VERSION : 0.1
   VAR_IN_OUT
      commands : "Linked List: Method Interface: Search";
      list : "Linked List: List";
   END_VAR
   VAR_TEMP
      clear_commands : "Linked List: Method Interface: Search";
      found : Bool;
      pointer_list : DInt;
   END_VAR
   VAR CONSTANT
      no_error : String := 'no error';
      searched_empty_list : String := 'searched empty list';
   END_VAR
BEGIN
   REGION "EXIT CONDITION: SEARCHED EMPTY LIST"
       IF "Linked List: Private: Is Empty"(#list) THEN
           #commands := #clear_commands;
           #commands.out.not_found := TRUE;
           #commands.out.error := TRUE;
           #commands.out.error_message := #searched_empty_list;
           RETURN;
       END_IF;
   END_REGION

   REGION "SEARCH"
       FOR #pointer_list := 0 TO "LINKED_LIST_LENGTH" DO
           IF #list.me[#pointer_list].data = #commands.in.data THEN
               #found := TRUE;
               EXIT;
           END_IF;
       END_FOR;
   END_REGION

   REGION "FOUND"
       IF #found THEN
           #commands := #clear_commands;
           #commands.out.done := TRUE;
           #commands.out.found := TRUE;
           #commands.out.returned_node := #list.me[#pointer_list];
           #commands.out.error_message := #no_error;
           RETURN;
       END_IF;
   END_REGION

   REGION "NOT FOUND"
       IF NOT #found THEN
           #commands := #clear_commands;
           #commands.out.done := TRUE;
           #commands.out.not_found := TRUE;
           RETURN;
       END_IF;
   END_REGION
END_FUNCTION

FUNCTION "Linked List: Display" : Void   // FC172, SCL
{ S7_Optimized_Access := 'TRUE' }
VERSION : 0.1
   VAR_IN_OUT
      commands : "Linked List: Method Interface: Display";
      list : "Linked List: List";
   END_VAR
   VAR_TEMP
      clear_commands : "Linked List: Method Interface: Display";
   END_VAR
BEGIN
   #commands := #clear_commands;
   #commands.out.list := #list;
   #commands.out.done := TRUE;
END_FUNCTION

FUNCTION "Linked List: Insert" : Void   // FC173, SCL
{ S7_Optimized_Access := 'TRUE' }
VERSION : 0.1
   VAR_INPUT
      terminal_behavior : String;
   END_VAR
   VAR_IN_OUT
      commands : "Linked List: Method Interface: Insert";
      list : "Linked List: List";
   END_VAR
   VAR_TEMP
      clear_commands : "Linked List: Method Interface: Insert";
      current : "Linked List: Node";
      next_empty_node_index : DInt;
      previous : "Linked List: Node";
      next : "Linked List: Node";
   END_VAR
   VAR CONSTANT
      no_error : String := 'no error';
      inserted_into_full : String := 'attempted to insert into full list. delete a node and try again.';
      appended_as_head : String := 'appended as head of list';
   END_VAR
BEGIN
   REGION "EXIT CONDITION: INSERTED INTO FULL LIST"
       IF "Linked List: Private: Is Full"(#list) THEN
           #commands := #clear_commands;
           #commands.out.error := TRUE;
           #commands.out.error_message := #inserted_into_full;
           RETURN;
       END_IF;
   END_REGION

   REGION "EXIT CONDITION: INSERTED INTO EMPTY LIST"
       IF "Linked List: Private: Is Empty"(#list) THEN
           "Linked List: Private: Head an Empty List"(data := #commands.in.data,
                                                      terminal_behavior := #terminal_behavior,
                                                      list := #list);
           #commands := #clear_commands;
           #commands.out.error := TRUE;
           #commands.out.error_message := #appended_as_head;
           RETURN;
       END_IF;
   END_REGION

   REGION "GET INDEX OF NEXT EMPTY NODE"
       #next_empty_node_index := "Linked List: Private: Next Empty Node"(#list);
   END_REGION

   REGION "PREVIOUS, CURRENT, AND NEXT NODES"
       #current := #commands.in.target_node;
       #previous := "Linked List: Private: Get Previous"(current := #current,
                                                         list := #list);
       #next := #current;
   END_REGION

   REGION "INSERT BEFORE TARGET NODE"
       // new node's data becomes command data
       #list.me[#next_empty_node_index].data := #commands.in.data;
       // new node's key becomes array index
       #list.me[#next_empty_node_index].meta.key := #next_empty_node_index;
       // shorten name for indexing
       #current := #list.me[#next_empty_node_index];
       // insert
       IF NOT #next.meta.is_head THEN
           "Linked List: Private: After"(node := #list.me[#current.meta.key],
                                         previous_node := #list.me[#previous.meta.key]);
       END_IF;
       "Linked List: Private: Before"(next_node := #list.me[#next.meta.key],
                                      node := #list.me[#current.meta.key]);
   END_REGION

   REGION "COMMANDS OUT"
       #commands := #clear_commands;
       #commands.out.done := TRUE;
       #commands.out.error_message := #no_error;
   END_REGION
END_FUNCTION

FUNCTION "Linked List: Reverse" : Void   // FC174, SCL
{ S7_Optimized_Access := 'TRUE' }
VERSION : 0.1
   VAR_IN_OUT
      commands : "Linked List: Method Interface: Reverse";
      list : "Linked List: List";
   END_VAR
   VAR_TEMP
      clear_commands : "Linked List: Method Interface: Reverse";
      current : "Linked List: Node";
      next : "Linked List: Node";
      previous : "Linked List: Node";
      null_node : "Linked List: Node";
   END_VAR
   VAR CONSTANT
      no_error : String := 'no error';
      reversed_empty_list : String := 'reversed empty list';
   END_VAR
BEGIN
   IF "Linked List: Private: Is Empty"(#list) THEN
       #commands := #clear_commands;
       #commands.out.error := TRUE;
       #commands.out.error_message := #reversed_empty_list;
       RETURN;
   END_IF;

   "Linked List: Private: Clear Node"(#null_node);
   #previous := #null_node;
   #current := "Linked List: Private: Get Head"(#list);
   #list.me[#current.meta.key].meta.is_head := FALSE;
   #list.me[#current.meta.key].meta.is_tail := TRUE;
   WHILE #current.meta.next <> "NULL_TOKEN" DO
       #next := #list.me[#current.meta.next];
       #list.me[#current.meta.key].meta.next := #previous.meta.key;
       #previous := #current;
       #current := #next;
       #list.me[#current.meta.key].meta.is_head := FALSE;
       #list.me[#current.meta.key].meta.is_tail := FALSE;
   END_WHILE;
   #list.me[#current.meta.key].meta.next := #previous.meta.key;
   #list.me[#current.meta.key].meta.is_head := TRUE;
   #list.me[#current.meta.key].meta.is_tail := FALSE;

   #commands := #clear_commands;
   #commands.out.done := TRUE;
   #commands.out.error_message := #no_error;
END_FUNCTION

FUNCTION "Linked List: Reset" : Void   // FC175, SCL
{ S7_Optimized_Access := 'TRUE' }
VERSION : 0.1
   VAR_IN_OUT
      commands : "Linked List: Method Interface: Reset";
      list : "Linked List: List";
   END_VAR
   VAR_TEMP
      blank_node : "Linked List: Node";
      list_pointer : DInt;
      clear_commands : "Linked List: Method Interface: Reset";
   END_VAR
BEGIN
   FOR #list_pointer := 0 TO "LINKED_LIST_LENGTH" DO
       "Linked List: Private: Clear Node"(#list.me[#list_pointer]);
   END_FOR;
   #commands := #clear_commands;
   #commands.out.done := TRUE;
END_FUNCTION

// folder: OBs

ORGANIZATION_BLOCK "Rack or station failure"   // OB86, LAD, RackStationFailure
{ S7_Optimized_Access := 'TRUE' }
VERSION : 0.1
   VAR_INPUT
      LADDR : Hw_Device;   // Hardware identifier
      Event_Class : Byte;   // Event class
      Fault_ID : Byte;   // Fault identifier
   END_VAR
BEGIN
END_ORGANIZATION_BLOCK

ORGANIZATION_BLOCK "Startup"   // OB100, LAD, Startup
TITLE = "Complete Restart"
{ S7_Optimized_Access := 'TRUE' }
VERSION : 0.1
   VAR_INPUT
      LostRetentive : Bool;   // True if retentive data are lost
      LostRTC : Bool;   // True if date and time are lost
   END_VAR
   VAR CONSTANT
      ALLOTTED : Real := 1800.0;
      CRITICAL : Real := 300.0;
   END_VAR
BEGIN

REGION Network 1
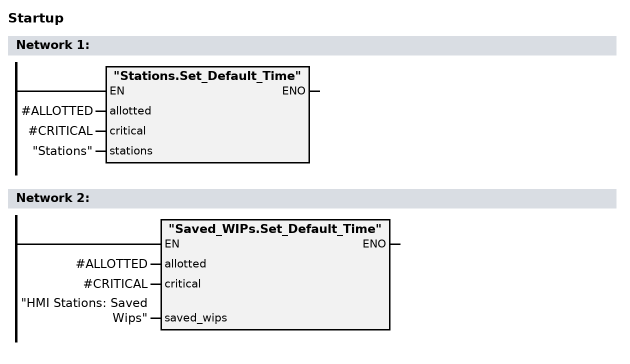
   RUNG wire#powerrail
      "Stations.Set_Default_Time"(allotted := #ALLOTTED, critical := #CRITICAL, stations := "Stations")
   END_RUNG
   // the same network as SCL:
   "Stations.Set_Default_Time"(allotted := #ALLOTTED, critical := #CRITICAL, stations := "Stations");
END_REGION

REGION Network 2
   RUNG wire#powerrail
      "Saved_WIPs.Set_Default_Time"(allotted := #ALLOTTED, critical := #CRITICAL, saved_wips := "HMI Stations: Saved Wips")
   END_RUNG
   // the same network as SCL:
   "Saved_WIPs.Set_Default_Time"(allotted := #ALLOTTED,
                           critical := #CRITICAL,
                           saved_wips := "HMI Stations: Saved Wips");
END_REGION
END_ORGANIZATION_BLOCK

ORGANIZATION_BLOCK "Programming error"   // OB121, LAD, ProgrammingError
{ S7_Optimized_Access := 'TRUE' }
VERSION : 0.1
   VAR_INPUT
      BlockNr : UInt;   // Number of causing block
      Reaction : USInt;   // 0:ignore, 1:substitute, 2:skip
      Fault_ID : Byte;   // Fault identifier
      BlockType : USInt;   // 16#01:OB, 16#02:FC, 16#03:FB, 16#04:SFC, 16#05:SFB, 16#06:DB: Type of block causing the error
      Area : USInt;   // Area where the error occured
      DBNr : DB_ANY;   // DB number if Area = DB or DI
      Csg_OBNr : OB_Any;   // Number of OB causing the error
      Csg_Prio : USInt;   // Priority of OB causing the error
      Width : USInt;   // 0:bit, 1:byte, 2:word, 3:dword, 4:lword
   END_VAR
BEGIN
END_ORGANIZATION_BLOCK

ORGANIZATION_BLOCK "IO access error"   // OB122, LAD, IOAccessError
{ S7_Optimized_Access := 'TRUE' }
VERSION : 0.1
   VAR_INPUT
      BlockNr : UInt;   // Number of causing block
      Reaction : USInt;   // 0:ignore, 1:substitute, 2:skip
      Fault_ID : Byte;   // 16#42:reading, 16#43:writing
      BlockType : USInt;   // 16#01:OB, 16#02:FC, 16#03:FB, 16#04:SFC, 16#05:SFB, 16#06:DB: Type of block causing the error
      Area : USInt;   // 16#81:I, 16#82:Q: IO area where the IOaccess error occured
      DBNr : DB_ANY;   // Reserved for system
      Csg_OBNr : OB_Any;   // Number of OB causing the error
      Csg_Prio : USInt;   // Priority of OB causing the error
      Width : USInt;   // 0:bit, 1:byte, 2:word, 3:dword, 4:lword
   END_VAR
BEGIN
END_ORGANIZATION_BLOCK

// folder: Order/States

FUNCTION_BLOCK "Order_State"   // FB2, SCL
{ S7_Optimized_Access := 'TRUE' }
VERSION : 0.1
   VAR_INPUT
      part_number_library : "Recipe: PN Text Library";
   END_VAR
   VAR_IN_OUT
      stations : "Station: All Stations";
   END_VAR
   VAR_TEMP
      station_pointer : Int;
      button_pointer : Int;
      station : "Station: Single Station";
   END_VAR
BEGIN
   REGION "FOR EACH STATION"
       FOR #station_pointer := 0 TO "STATION_COUNT" DO

           REGION "POPULATE CURRENT STATION"
               #station := #stations.stn[#station_pointer];
           END_REGION

           REGION "SET TO IDLE ON WIP SWAP"
               IF #station.flags.wipSwapped THEN
                   CONTINUE;
               END_IF;
           END_REGION

           REGION "FOR EACH BUTTON"
               FOR #button_pointer := 0 TO "BUTTON_COUNT" DO

                   REGION "INITIALIZE STATE"
                       "Order_State.Initialize_State"(newParams := #station.wipCmpts.flags.new_part_number,
                                                      pnGood := #station.wipCmpts.flags.part_number_good[#button_pointer],
                                                      state := #station.wipCmpts.orderState[#button_pointer]);
                   END_REGION

                   REGION "ENTER IDLE"
                       "Order_State.Enter_Idle"(part_button_falling_edge := #station.wipCmpts.kp8Logical.falling.btn[#button_pointer],
                                                state := #station.wipCmpts.orderState[#button_pointer]);
                   END_REGION

                   REGION "ENTER REQUESTED"
                       "Order_State.Enter_Requested"(btnRising := #station.wipCmpts.kp8Logical.rising.btn[#button_pointer],
                                                     state := #station.wipCmpts.orderState[#button_pointer]);
                   END_REGION

                   REGION "ENTER REQUESTED CRITICAL"
                       "Order_State.Enter_Requested_Critical"(timerVal := #station.wipCmpts.timers.remaining[#button_pointer],
                                                              state := #station.wipCmpts.orderState[#button_pointer]);
                   END_REGION

                   REGION "ENTER REQUESTED EXPIRED"
                       "Order_State.Enter_Requested_Expired"(timerVal := #station.wipCmpts.timers.remaining[#button_pointer],
                                                             state := #station.wipCmpts.orderState[#button_pointer]);
                   END_REGION

                   REGION "SAVE CURRENT STATION"
                       #stations.stn[#station_pointer] := #station;
                   END_REGION

               END_FOR;
           END_REGION

       END_FOR;
   END_REGION
END_FUNCTION_BLOCK

FUNCTION "Order_State.Enter_Idle" : Void   // FC6, SCL
{ S7_Optimized_Access := 'TRUE' }
VERSION : 0.1
   VAR_INPUT
      part_button_falling_edge : Bool;
   END_VAR
   VAR_IN_OUT
      state : Int;
   END_VAR
BEGIN
   IF #part_button_falling_edge THEN
       #state := "IDLE";
       RETURN;
   END_IF;
END_FUNCTION

FUNCTION "Order_State.Enter_Requested" : Void   // FC7, SCL
{ S7_Optimized_Access := 'TRUE' }
VERSION : 0.1
   VAR_INPUT
      btnRising : Bool;
   END_VAR
   VAR_IN_OUT
      state : Int;
   END_VAR
BEGIN
   IF #state = "IDLE" THEN
       IF #btnRising THEN
           #state := "REQUESTED";
       END_IF;
   END_IF;
END_FUNCTION

FUNCTION "Order_State.Initialize_State" : Void   // FC10, SCL
{ S7_Optimized_Access := 'TRUE' }
VERSION : 0.1
   VAR_INPUT
      newParams : Bool;
      pnGood : Bool;
   END_VAR
   VAR_IN_OUT
      state : Int;
   END_VAR
BEGIN
   REGION "ON NEW PARAMETERS"
       IF #newParams THEN
           #state := BOOL_TO_INT(#pnGood);
       END_IF;
   END_REGION
END_FUNCTION

FUNCTION "Order_State.Enter_Requested_Critical" : Void   // FC16, SCL
{ S7_Optimized_Access := 'TRUE' }
VERSION : 0.1
   VAR_INPUT
      timerVal : Real;
   END_VAR
   VAR_IN_OUT
      state : Int;
   END_VAR
   VAR_TEMP
      temp : Real;
   END_VAR
BEGIN
   IF #state = "REQUESTED" THEN
       IF #timerVal > 0.0 AND #timerVal <= "DEFAULT_CRITICAL_TIME" THEN
           #state := "REQUESTED_CRITICAL";
       END_IF;
   END_IF;
END_FUNCTION

FUNCTION "Order_State.Enter_Requested_Expired" : Void   // FC17, SCL
{ S7_Optimized_Access := 'TRUE' }
VERSION : 0.1
   VAR_INPUT
      timerVal : Real;
   END_VAR
   VAR_IN_OUT
      state : Int;
   END_VAR
BEGIN
   IF #state = "REQUESTED_CRITICAL" THEN
       IF #timerVal <= -0.001 THEN
           #state := "REQUESTED_EXPIRED";
       END_IF;
   END_IF;
END_FUNCTION

FUNCTION "Order_State.Enter_Ordered" : Void   // FC297, SCL
{ S7_Optimized_Access := 'TRUE' }
VERSION : 0.1
   VAR_INPUT
      address : DInt;
   END_VAR
   VAR_IN_OUT
      stations : "Station: All Stations";
   END_VAR
BEGIN
   "Order_State.Set_State_by_Address"(address := #address,
                                      state := "ORDERED",
                                      stations := #stations);
END_FUNCTION

FUNCTION "Order_State.Enter_Acknowledged" : Void   // FC301, SCL
{ S7_Optimized_Access := 'TRUE' }
VERSION : 0.1
   VAR_INPUT
      address : DInt;
   END_VAR
   VAR_IN_OUT
      stations : "Station: All Stations";
   END_VAR
BEGIN
   "Order_State.Set_State_by_Address"(address := #address,
                                      state := "ACKNOWLEGED",
                                      stations := #stations);
END_FUNCTION

FUNCTION "Order_State.Set_State_by_Address" : Void   // FC302, SCL
{ S7_Optimized_Access := 'TRUE' }
VERSION : 0.1
   VAR_INPUT
      address : DInt;
      state : Int;
   END_VAR
   VAR_IN_OUT
      stations : "Station: All Stations";
   END_VAR
   VAR_TEMP
      _p_button : DInt;
      _p_station : DInt;
      _p_wip : DInt;
   END_VAR
BEGIN
   #_p_button := "Address.Get_Button"(#address);
   #_p_station := "Address.Get_Station"(#address);
   #_p_wip := "Address.Get_Wip"(#address);
   #stations.stn[#_p_station].wipCmpts.orderState[#_p_button] := #state;
END_FUNCTION

FUNCTION "Order_State.Swap_WIP_States" : Void   // FC317, SCL
{ S7_Optimized_Access := 'TRUE' }
VERSION : 0.1
   VAR_IN_OUT
      station : "Station: Single Station";
   END_VAR
   VAR_TEMP
      _length : Int;
      _button_pointer : Int;
   END_VAR
BEGIN
   #_length := UDINT_TO_INT("Array.Any.Length"(#station.wipCmpts.pnCode)) - 1;
   FOR #_button_pointer := 0 TO #_length DO
       IF #station.wipCmpts.pnCode[#_button_pointer] <= 0 THEN
           #station.wipCmpts.orderState[#_button_pointer] := 0;
           CONTINUE;
       END_IF;
       IF #station.wipCmpts.orderState[#_button_pointer] <> 0 THEN
           CONTINUE;
       END_IF;
       #station.wipCmpts.orderState[#_button_pointer] := "IDLE";
   END_FOR;
END_FUNCTION

// folder: Order/Timers

FUNCTION_BLOCK "Order Timer"   // FB6, SCL
{ S7_Optimized_Access := 'TRUE' }
VERSION : 0.1
   VAR_INPUT
      pnLib : "Recipe: PN Text Library";
   END_VAR
   VAR_IN_OUT
      stns : "Station: All Stations";
   END_VAR
   VAR
      rt : "Runtime Data";
   END_VAR
   VAR_TEMP
      pStn : Int;
      pBtn : Int;
   END_VAR
BEGIN
   REGION "RUNTIME CALL"
       #rt.elapsed := RUNTIME(#rt.mem);
       #rt.asReal := LREAL_TO_REAL(#rt.elapsed);
   END_REGION

   REGION "FOR EACH STATION"
       FOR #pStn := 0 TO "STATION_COUNT" DO

           REGION "FOR EACH BUTTON"
               FOR #pBtn := 0 TO "BUTTON_COUNT" DO

                   REGION "INITIALIZE TIMERS"
                       "Order Timer: Initialize"(pnLib := #pnLib,
                                                 pBtn := #pBtn,
                                                 stn := #stns.stn[#pStn]);
                   END_REGION

                   REGION "EXECUTE TIMERS"
                       "Order Timer: Timer Execution"(elapsedTime := #rt.asReal,
                                                      pBtn := #pBtn,
                                                      stn:=#stns.stn[#pStn],
                                                      timers := #stns.stn[#pStn].wipCmpts.timers);
                   END_REGION

               END_FOR;
           END_REGION

       END_FOR;
   END_REGION
END_FUNCTION_BLOCK

FUNCTION "Order Timer: Initialize" : Void   // FC8, SCL
{ S7_Optimized_Access := 'TRUE' }
VERSION : 0.1
   VAR_INPUT
      pnLib : "Recipe: PN Text Library";
      pBtn : Int;
   END_VAR
   VAR_IN_OUT
      stn : "Station: Single Station";
   END_VAR
   VAR_TEMP
      pnGood : Bool;
      default : Bool;
      clear : Bool;
   END_VAR
BEGIN
   REGION "ON PN CHANGE"
       IF #stn.wipCmpts.flags.new_part_number THEN

           REGION "INITIALIZE TO DEFAULT"

               REGION "EXECUTION VALIDATION"
                   #default := "Order Timer: Set to Default Check"(pnGood := #stn.wipCmpts.flags.part_number_good[#pBtn],
                                                                   inSettingsScreen := #stn.wipCmpts.flags.in_settings_screen,
                                                                   timerReset := #stn.wipCmpts.flags.reset_timer[#pBtn]);
               END_REGION

               REGION "ON VALIDATION"
                   IF #default THEN

                       REGION "SET DEFAULT TIME VALUE"
                           #stn.wipCmpts.timers.ptAllotted[#pBtn] := "DEFAULT_TOTAL_TIME";
                           #stn.wipCmpts.timers.ptCritical[#pBtn] := "DEFAULT_CRITICAL_TIME";
                       END_REGION

                   END_IF;
               END_REGION

           END_REGION

           REGION "INITIALIZE TO ZERO"

               REGION "EXECUTION VALIDATION"
                   #clear := "Order Timer: Set to Zero Check"(pnGood := #stn.wipCmpts.flags.part_number_good[#pBtn],
                                                              inSettingsScreen := #stn.wipCmpts.flags.in_settings_screen,
                                                              timerReset := #stn.wipCmpts.flags.reset_timer[#pBtn]);
               END_REGION

               REGION "ON VALIDATION"
                   IF #clear THEN

                       REGION "SET DEFAULT TIME VALUE"
                           #stn.wipCmpts.timers.ptAllotted[#pBtn] := 0.0;
                           #stn.wipCmpts.timers.ptCritical[#pBtn] := 0.0;
                       END_REGION

                   END_IF;
               END_REGION

           END_REGION

       END_IF;
   END_REGION
END_FUNCTION

FUNCTION "Order Timer: Timer Execution" : Void   // FC11, SCL
{ S7_Optimized_Access := 'TRUE' }
VERSION : 0.1
   VAR_INPUT
      elapsedTime : Real;
      pBtn : Int;
      stn : "Station: Single Station";
   END_VAR
   VAR_IN_OUT
      timers : "Request_Timers.UDT";
   END_VAR
BEGIN
   REGION "RUN CONDITIONS"
       CASE #stn.wipCmpts.orderState[#pBtn] OF

           "RESET", "IDLE":
               IF #stn.flags.stateTransition[#pBtn] THEN
                   #timers.elapsed[#pBtn] := 0.0;
                   #timers.remaining[#pBtn] := 0.0;
               END_IF;

           "REQUESTED".."ACKNOWLEDGED_EXPIRED":
               #timers.elapsed[#pBtn] += #elapsedTime;
               #timers.remaining[#pBtn] := #timers.ptAllotted[#pBtn] - #timers.elapsed[#pBtn];

           ELSE:
               ;

       END_CASE;
   END_REGION
END_FUNCTION

FUNCTION "Order Timer: Set to Default Check" : Bool   // FC12, SCL
{ S7_Optimized_Access := 'TRUE' }
VERSION : 0.1
   VAR_INPUT
      pnGood : Bool;
      inSettingsScreen : Bool;
      timerReset : Bool;
   END_VAR
   VAR_TEMP
      ret : Bool;
   END_VAR
BEGIN
   REGION "ON VALID PN"
       #ret := #pnGood;
   END_REGION

   REGION "NOT WHILE IN SETTINGS SCREEN"
       IF #inSettingsScreen THEN
           #ret := FALSE;
       END_IF;
   END_REGION

   REGION "ON RESET REQUEST"
       #ret := #timerReset OR #ret;
   END_REGION

   REGION "RETURN"
       #"Order Timer: Set to Default Check" := #ret;
   END_REGION
END_FUNCTION

FUNCTION "Order Timer: Set to Zero Check" : Bool   // FC15, SCL
{ S7_Optimized_Access := 'TRUE' }
VERSION : 0.1
   VAR_INPUT
      pnGood : Bool;
      inSettingsScreen : Bool;
      timerReset : Bool;
   END_VAR
   VAR_TEMP
      ret : Bool;
   END_VAR
BEGIN
   REGION "ON VALID PN"
       #ret := NOT #pnGood;
   END_REGION

   REGION "NOT WHILE IN SETTINGS SCREEN"
       IF #inSettingsScreen THEN
           #ret := FALSE;
       END_IF;
   END_REGION

   REGION "ON RESET REQUEST"
       #ret := #timerReset OR #ret;
   END_REGION

   REGION "RETURN"
       #"Order Timer: Set to Zero Check" := #ret;
   END_REGION
END_FUNCTION

// folder: Part Request

FUNCTION_BLOCK "Part Request"   // FB7, SCL
{ S7_Optimized_Access := 'TRUE' }
VERSION : 0.1
   VAR_INPUT
      stns : "Station: All Stations";
      savedWips : "Recipe: HMI Stations Saved Wips";
      pnLib : "Recipe: PN Text Library";
   END_VAR
   VAR_IN_OUT
      dataTable : "Part Request Data";
   END_VAR
   VAR RETAIN
      pDataRow : Int;
   END_VAR
   VAR_TEMP
      address : DInt;
      addRequest : Bool;
      inTable : DInt;
      pStn : Int;
      pBtn : Int;
      pWip : Int;
      pRqstsRow : Int;
      removeRequest : Bool;
   END_VAR
BEGIN
   REGION "FOR EACH STATION"
       FOR #pStn := 0 TO "STATION_COUNT" DO

           REGION "FOR EACH BUTTON"
               FOR #pBtn := 0 TO "BUTTON_COUNT" DO

                   REGION "NEXT BUTTON ON NO TRANSITION"
                       IF NOT #stns.stn[#pStn].flags.stateTransition[#pBtn] THEN
                           CONTINUE;
                       END_IF;
                   END_REGION

                   REGION "GET ADDRESS"
                       #pWip := DINT_TO_INT(#stns.stn[#pStn].wipData.index);
                       #address := "Address.Set_Address"(pStn := #pStn, pBtn := #pBtn, pWip := #pWip);
                   END_REGION

                   REGION "CHECK FOR ENTRY IN DATA TABLE"
                       #inTable := "Part Request: Address in Table"(address := #address,
                                                                    table := #dataTable);
                   END_REGION

                   REGION "ADD"

                       REGION "VALIDATE CONDITIONS"
                           #addRequest := "Part Request: Validate Add"(inTable := #inTable,
                                                                       orderState := #stns.stn[#pStn].wipCmpts.orderState[#pBtn]);
                       END_REGION

                       REGION "EXECUTE"
                           IF #addRequest THEN
                               #addRequest := FALSE;
                               #dataTable.row[#pDataRow] := #address;
                               "Row Pointer: Roll Over"(limit := "partReqDataRowCount",
                                                        "pointer" := #pDataRow);
                           END_IF;
                       END_REGION

                   END_REGION

                   REGION "REMOVE SINGLE STATION"

                       REGION "VALIDATE CONDITIONS: SINGLE"
                           #removeRequest := "Part Request: Validate Remove: Single"(inTable := #inTable,
                                                                                     orderState := #stns.stn[#pStn].wipCmpts.orderState[#pBtn]);
                       END_REGION

                       REGION "EXECUTE"
                           IF #removeRequest THEN
                               #removeRequest := FALSE;
                               #dataTable.row[#inTable] := -1;
                               "Part Request: Collapse Table"(#dataTable);
                               "Row Pointer: Post Collapse"(dataTable := #dataTable,
                                                            pDataRow := #pDataRow);
                           END_IF;
                       END_REGION

                   END_REGION

               END_FOR;
           END_REGION

       END_FOR;
   END_REGION
END_FUNCTION_BLOCK

FUNCTION "Part Request: Address in Table" : DInt   // FC27, SCL
{ S7_Optimized_Access := 'TRUE' }
VERSION : 0.1
   VAR_INPUT
      address : DInt;
      table : "Part Request Data";
   END_VAR
   VAR_TEMP
      _i : DInt;
      _length : DInt;
   END_VAR
BEGIN
   #_length := UDINT_TO_DINT("Array.Any.Length"(#table.row)) - 1;
   FOR #_i := 0 TO #_length DO
       IF #table.row[#_i] = #address THEN
           #"Part Request: Address in Table" := #_i;
           RETURN;
       END_IF;
   END_FOR;
   #"Part Request: Address in Table" := "NULL_TOKEN";
END_FUNCTION

FUNCTION "Part Request: Validate Add" : Bool   // FC30, SCL
{ S7_Optimized_Access := 'TRUE' }
VERSION : 0.1
   VAR_INPUT
      inTable : DInt;
      orderState : Int;
   END_VAR
   VAR_TEMP
      ret : Bool;
   END_VAR
BEGIN
   IF #inTable = -1 THEN
       CASE #orderState OF
           "IDLE",
           "REQUESTED_CRITICAL", "REQUESTED_EXPIRED",
           "ORDERED", "ORDERED_CRITICAL", "ORDERED_EXPIRED",
           "ACKNOWLEGED", "ACKNOWLEDGED_CRITICAL", "ACKNOWLEDGED_EXPIRED":
               #ret := FALSE;
           "REQUESTED":
               #ret := TRUE;
       END_CASE;
   END_IF;
   #"Part Request: Validate Add" := #ret;
END_FUNCTION

FUNCTION "Part Request: Validate Remove: Single" : Bool   // FC41, SCL
{ S7_Optimized_Access := 'TRUE' }
VERSION : 0.1
   VAR_INPUT
      inTable : DInt;
      orderState : Int;
   END_VAR
   VAR_TEMP
      ret : Bool;
   END_VAR
BEGIN
   IF #inTable <> -1 THEN
       CASE #orderState OF
           "REQUESTED", "REQUESTED_CRITICAL", "REQUESTED_EXPIRED",
           "ORDERED", "ORDERED_CRITICAL", "ORDERED_EXPIRED",
           "ACKNOWLEGED", "ACKNOWLEDGED_CRITICAL", "ACKNOWLEDGED_EXPIRED":
               #ret := FALSE;
           "IDLE":
               #ret := TRUE;
       END_CASE;
   END_IF;
   #"Part Request: Validate Remove: Single" := #ret;
END_FUNCTION

FUNCTION "Part Request: Clear Data Table" : Void   // FC48, SCL
{ S7_Optimized_Access := 'TRUE' }
VERSION : 0.1
   VAR_IN_OUT
      dataTable : "Part Request Data";
   END_VAR
   VAR_TEMP
      pRow : Int;
   END_VAR
   VAR CONSTANT
      clearRow : DInt := -1;
   END_VAR
BEGIN
   FOR #pRow := 0 TO "partReqDataRowCount" DO
       #dataTable.row[#pRow] := #clearRow;
   END_FOR;
END_FUNCTION

FUNCTION "Part Request: Collapse Table" : Void   // FC55, SCL
{ S7_Optimized_Access := 'TRUE' }
VERSION : 0.1
   VAR_IN_OUT
      dataTable : "Part Request Data";
   END_VAR
   VAR_TEMP
      pRow : Int;
      pScan : Int;
   END_VAR
BEGIN
   FOR #pRow := 0 TO "partReqDataRowCount" DO
       #pScan := 1;
       IF #dataTable.row[#pRow] <= -1 THEN
           WHILE #dataTable.row[#pRow + #pScan] <= -1 AND #pRow + #pScan < "partReqDataRowCount" DO
               #pScan += 1;
           END_WHILE;
           #dataTable.row[#pRow] := #dataTable.row[#pRow + #pScan];
           #dataTable.row[#pRow + #pScan] := -1;
           IF #pRow + #pScan = "partReqDataRowCount" THEN
               RETURN;
           END_IF;
       END_IF;
   END_FOR;
END_FUNCTION

FUNCTION "Part Request: Validate Remove: WIP" : Bool   // FC89, SCL
{ S7_Optimized_Access := 'TRUE' }
VERSION : 0.1
   VAR_INPUT
      inTable : DInt;
      clearWipRequest : Bool;
   END_VAR
   VAR_TEMP
      ret : Bool;
   END_VAR
BEGIN
   IF #inTable <> -1 THEN
       #ret := #clearWipRequest;
   END_IF;

   #"Part Request: Validate Remove: WIP" := #ret;
END_FUNCTION

// folder: Request_Table

FUNCTION_BLOCK "Request_Table.Row_Selection"   // FB61, SCL
{ S7_Optimized_Access := 'TRUE' }
VERSION : 0.1
   VAR_INPUT
      request_table : "Part Call Screen";
   END_VAR
   VAR_IN_OUT
      barcode_data : "Barcode.UDT";
   END_VAR
   VAR
      last_selection : Int := -1;
   END_VAR
   VAR_TEMP
      _selected_row : Int;
   END_VAR
BEGIN
   #_selected_row := "Request_Table.Get_Selected_Row_Index"(#request_table);
   IF #_selected_row = "NULL_TOKEN" THEN
       #last_selection := #_selected_row;
       RETURN;
   END_IF;
   IF #_selected_row <> #last_selection THEN
       "Barcode.Load_Data"(address := #request_table.row[#_selected_row].address,
                           part_number := #request_table.row[#_selected_row].tfPartNumber.value,
                           barcode_data := #barcode_data);
   END_IF;
   #last_selection := #_selected_row;
END_FUNCTION_BLOCK

FUNCTION "Request_Table.Navigation_Animations" : Void   // FC18, SCL
{ S7_Optimized_Access := 'TRUE' }
VERSION : 0.1
   VAR_IN_OUT
      tableNav : "Nav Bar Data: PLC";
   END_VAR
   VAR_TEMP
      gray : USInt;
      green : USInt;
   END_VAR
BEGIN
   REGION "ANIMATE PART CALL NAV"

       REGION "COPY TO LOCAL"
           #gray := "GRAY_BACKGROUND";
           #green := "GREEN_LIGHT_BACKGROUND";
       END_REGION

       REGION "TOP"
           #tableNav.top.animate := "Bool.Animate"(true_color := #green,
                                                   false_color := #gray,
                                                   evaluation_signal := #tableNav.top.actuate);
       END_REGION

       REGION "PAGE UP"
           #tableNav.pageUp.animate := "Bool.Animate"(true_color := #green,
                                                      false_color := #gray,
                                                      evaluation_signal := #tableNav.pageUp.actuate);
       END_REGION

       REGION "LINE UP"
           #tableNav.lineUp.animate := "Bool.Animate"(true_color := #green,
                                                      false_color := #gray,
                                                      evaluation_signal := #tableNav.lineUp.actuate);
       END_REGION

       REGION "LINE DOWN"
           #tableNav.lineDown.animate := "Bool.Animate"(true_color := #green,
                                                        false_color := #gray,
                                                        evaluation_signal := #tableNav.lineDown.actuate);
       END_REGION

       REGION "PAGE DOWN"
           #tableNav.pageDown.animate := "Bool.Animate"(true_color := #green,
                                                        false_color := #gray,
                                                        evaluation_signal := #tableNav.pageDown.actuate);
       END_REGION

       REGION "BOTTOM"
           #tableNav.bottom.animate := "Bool.Animate"(true_color := #green,
                                                      false_color := #gray,
                                                      evaluation_signal := #tableNav.bottom.actuate);
       END_REGION

   END_REGION
END_FUNCTION

FUNCTION "Request_Table.State_to_Color" : Void   // FC22, SCL
{ S7_Optimized_Access := 'TRUE' }
VERSION : 0.1
   VAR_INPUT
      state : Int;
   END_VAR
   VAR_OUTPUT
      background : USInt;
      foreground : USInt;
   END_VAR
   VAR_TEMP
      bg : USInt;
      cBlue : USInt;
      cGrayLight : USInt;
      cGrayDark : USInt;
      cGreen : USInt;
      cInvisible : USInt;
      cRedSolid : USInt;
      cRedFlash : USInt;
      cWhite : USInt;
      fg : USInt;
   END_VAR
BEGIN
   #cBlue := "BLUE_LIGHT_BACKGROUND";
   #cGreen := "GREEN_LIGHT_BACKGROUND";
   #cInvisible := "INVISIBLE";
   #cRedSolid := "RED_LIGHT_BACKGROUND";
   #cRedFlash := "RED_LIGHT_FLASHING";
   #cGrayLight := "GRAY_BACKGROUND";
   #cGrayDark := "DISABLED";
   #cWhite := "WHITE_BACKGROUND";

   CASE #state OF
       0, "IDLE":
           #bg := #cInvisible;
           #fg := #cInvisible;
       "REQUESTED":
           #bg := #cGrayDark;
           #fg := #cGrayLight;
       "ACKNOWLEGED":
           #bg := #cGrayDark;
           #fg := "YELLOW_LIGHT_BACKGROUND";
       "REQUESTED_CRITICAL", "ORDERED_CRITICAL", "ACKNOWLEDGED_CRITICAL":
           #bg := #cGrayDark;
           #fg := #cRedSolid;
       "REQUESTED_EXPIRED", "ORDERED_EXPIRED", "ACKNOWLEDGED_EXPIRED":
           #bg := #cGrayDark;
           #fg := #cRedFlash;
       "ORDERED":
           #bg := #cGrayDark;
           #fg := #cBlue;
   END_CASE;

   #foreground := #fg;
   #background := #bg;
END_FUNCTION

FUNCTION "Request_Table.Get_States" : Int   // FC57, SCL
{ S7_Optimized_Access := 'TRUE' }
VERSION : 0.1
   VAR_INPUT
      address : DInt;
      stations : "Station: All Stations";
      saved_wips : "Recipe: HMI Stations Saved Wips";
   END_VAR
   VAR_TEMP
      _address_in_wip : Bool;
      _button_pointer : DInt;
      _saved_station_pointer : DInt;
      _station_pointer : DInt;
      _wip_pointer : DInt;
   END_VAR
BEGIN
   REGION "DECOMPOSE ADDRESS"
       #_button_pointer := "Address.Get_Button"(#address);
       #_station_pointer := "Address.Get_Station"(#address);
       #_wip_pointer := "Address.Get_Wip"(#address);
   END_REGION

   REGION "CHECK ADDRESS AGAINST STATION'S CURRENT WIP"
       #_address_in_wip := "Address in Loaded Wip"(pWip := #_wip_pointer,
                                                   stn := #stations.stn[#_station_pointer]);
   END_REGION

   REGION "ADDRESS IN WIP"
       IF #_address_in_wip THEN
           #"Request_Table.Get_States" := #stations.stn[#_station_pointer].wipCmpts.orderState[#_button_pointer];
           RETURN;
       END_IF;
   END_REGION

   REGION "ADDRESS NOT IN WIP"
       #_saved_station_pointer := "WIP.Global_Index_to_HMI_Station_Index"(global_index := DINT_TO_INT(#_station_pointer),
                                                                          saved_WIPs := #saved_wips);
       #"Request_Table.Get_States" := #saved_wips.stn[#_saved_station_pointer].wip[#_wip_pointer].orderState[#_button_pointer];
   END_REGION
END_FUNCTION

FUNCTION "Request_Table.Draw" : Void   // FC295, SCL
{ S7_Optimized_Access := 'TRUE' }
VERSION : 0.1
   VAR_INPUT
      pn_library : "Recipe: PN Text Library";
      row_indices : Array[*] of DInt;   // needs to be same length as request_table
      saved_wips : "Recipe: HMI Stations Saved Wips";
      stations : "Station: All Stations";
      table_data : "Part Request Data";
   END_VAR
   VAR_IN_OUT
      request_table : Array[*] of "Table Row";   // needs to be same length as row_indices
   END_VAR
   VAR_TEMP
      _length_indices : DInt;
      _length_table : DInt;
      _p_row_hmi : DInt;
      _p_row_data : DInt;
   END_VAR
BEGIN
   REGION "GET LENGTH"
       #_length_indices := UDINT_TO_DINT("Array.Any.Length"(#row_indices)) - 1;
       #_length_table := UDINT_TO_DINT("Array.Any.Length"(#request_table)) - 1;
   END_REGION


   REGION "EXIT ON MISMATCHED LENGTH"
       IF #_length_indices <> #_length_table THEN
           RETURN;
       END_IF;
   END_REGION


   REGION "DRAW HMI TABLE"
       FOR #_p_row_hmi := 0 TO #_length_table DO
           #_p_row_data := #row_indices[#_p_row_hmi];
           "Table_Row.Draw"(address := #table_data.row[#_p_row_data],
                            pn_library := #pn_library,
                            stations := #stations,
                            saved_wips := #saved_wips,
                            row_hmi := #request_table[#_p_row_hmi]);
       END_FOR;
   END_REGION
END_FUNCTION

FUNCTION "Request_Table.Get_Selected_Row_Index" : Int   // FC299, SCL
{ S7_Optimized_Access := 'TRUE' }
VERSION : 0.1
   VAR_INPUT
      request_table : "Part Call Screen";
   END_VAR
   VAR_TEMP
      _length : Int;
      _i : Int;
   END_VAR
BEGIN
   #_length := UDINT_TO_INT("Array.Any.Length"(#request_table.row)) - 1;
   FOR #_i := 0 TO #_length DO
       IF #request_table.row[#_i].pbSelection.actuate THEN
           #"Request_Table.Get_Selected_Row_Index" := #_i;
           RETURN;
       END_IF;
   END_FOR;
   #"Request_Table.Get_Selected_Row_Index" := "NULL_TOKEN";
   RETURN;
END_FUNCTION

// folder: Request_Timers

FUNCTION "Request_Timers.Set_Default_Time" : Void   // FC321, SCL
{ S7_Optimized_Access := 'TRUE' }
VERSION : 0.1
   VAR_INPUT
      allotted : Real;
      critical : Real;
   END_VAR
   VAR_IN_OUT
      wip_module : "WIP_Module.UDT";
   END_VAR
   VAR_TEMP
      _i : Int;
      _length : Int;
   END_VAR
BEGIN
   #_length := UDINT_TO_INT("Array.Any.Length"(#wip_module.pnCode)) - 1;
   FOR #_i := 0 TO #_length DO
       CASE #wip_module.pnCode[#_i] OF
           0, "NULL_TOKEN":
               CONTINUE;
           ELSE
               #wip_module.timers.ptAllotted[#_i] := #allotted;
               #wip_module.timers.ptCritical[#_i] := #critical;
       END_CASE;
   END_FOR;
END_FUNCTION

// folder: Stack_Light

FUNCTION "Stack_Light.Green" : Void   // FC325, SCL
{ S7_Optimized_Access := 'TRUE' }
VERSION : 0.1
   VAR_INPUT
      part_number : Int;
   END_VAR
   VAR_IN_OUT
      stack_light : DWord;
   END_VAR
   VAR CONSTANT
      GREEN_ON_00 : DWord := 16#0400_0000;
      GREEN_ON_01 : DWord := 16#2000_0000;
      GREEN_ON_02 : DWord := 16#0001_0000;
      GREEN_ON_03 : DWord := 16#0008_0000;
      GREEN_ON_04 : DWord := 16#0040_0000;
      GREEN_ON_05 : DWord := 16#0000_0200;
      PART_00 : Int := 7;
      PART_01 : Int := 3;
      PART_02 : Int := 6;
      PART_03 : Int := 2;
      PART_04 : Int := 5;
      PART_05 : Int := 1;
   END_VAR
BEGIN
   CASE #part_number OF
       #PART_00:
           #stack_light := #stack_light OR #GREEN_ON_00;
       #PART_01:
           #stack_light := #stack_light OR #GREEN_ON_01;
       #PART_02:
           #stack_light := #stack_light OR #GREEN_ON_02;
       #PART_03:
           #stack_light := #stack_light OR #GREEN_ON_03;
       #PART_04:
           #stack_light := #stack_light OR #GREEN_ON_04;
       #PART_05:
           #stack_light := #stack_light OR #GREEN_ON_05;
       ELSE
           ;
   END_CASE;
END_FUNCTION

FUNCTION "Stack_Light.State_to_Color" : Void   // FC326, SCL
{ S7_Optimized_Access := 'TRUE' }
VERSION : 0.1
   VAR_INPUT
      part_number : Int;
      state : Int;
   END_VAR
   VAR_IN_OUT
      stack_light : DWord;
   END_VAR
BEGIN
   CASE #state OF

       "NO_STATE", "RESET":
           "Stack_Light.Off"(part_number := #part_number,
                             stack_light := #stack_light);

       "IDLE":
           "Stack_Light.Off"(part_number := #part_number,
                             stack_light := #stack_light);
           "Stack_Light.Green"(part_number := #part_number,
                               stack_light := #stack_light);

       "REQUESTED", "ORDERED", "ACKNOWLEGED":
           "Stack_Light.Off"(part_number := #part_number,
                             stack_light := #stack_light);
           "Stack_Light.Yellow"(part_number := #part_number,
                                stack_light := #stack_light);

       "REQUESTED_CRITICAL", "ORDERED_CRITICAL", "ACKNOWLEDGED_CRITICAL":
           "Stack_Light.Off"(part_number := #part_number,
                             stack_light := #stack_light);
           "Stack_Light.Red"(part_number := #part_number,
                             stack_light := #stack_light);

       "REQUESTED_EXPIRED", "ORDERED_EXPIRED", "ACKNOWLEDGED_EXPIRED":
           "Stack_Light.Off"(part_number := #part_number,
                             stack_light := #stack_light);
           "Stack_Light.Flash_Red"(part_number := #part_number,
                                   animator := "Clock_1.25Hz",
                                   stack_light := #stack_light);

       ELSE
           ;

   END_CASE;
END_FUNCTION

FUNCTION "Stack_Light.Animate_All_Stations" : Void   // FC327, SCL
{ S7_Optimized_Access := 'TRUE' }
VERSION : 0.1
   VAR_IN_OUT
      stations : "Station: All Stations";
   END_VAR
   VAR_TEMP
      _button_count : Int;
      _button_pointer : Int;
      _stack_light : DWord;
      _station_count : Int;
      _station_pointer : Int;
   END_VAR
BEGIN
   #_station_count := UDINT_TO_INT("Array.Any.Length"(#stations.stn)) - 1;
   #_button_count := UDINT_TO_INT("Array.Any.Length"(#stations.stn[0].wipCmpts.orderState)) - 1;

   REGION "LOOP THROUGH STATIONS"
       FOR #_station_pointer := 0 TO #_station_count DO

           REGION "LOOP THROUGH BUTTONS"
               FOR #_button_pointer := 0 TO #_button_count DO

                   #_stack_light := #stations.stn[#_station_pointer].wipCmpts.ioData.stkLight;
                   "Stack_Light.State_to_Color"(part_number := #_button_pointer,
                                                state := #stations.stn[#_station_pointer].wipCmpts.orderState[#_button_pointer],
                                                stack_light := #_stack_light);
                   #stations.stn[#_station_pointer].wipCmpts.ioData.stkLight := #_stack_light;

               END_FOR;
           END_REGION

       END_FOR;
   END_REGION
END_FUNCTION

FUNCTION "Stack_Light.Flash_Red" : Void   // FC328, SCL
{ S7_Optimized_Access := 'TRUE' }
VERSION : 0.1
   VAR_INPUT
      part_number : Int;
      animator : Bool;
   END_VAR
   VAR_IN_OUT
      stack_light : DWord;
   END_VAR
   VAR CONSTANT
      RED_ON_00 : DWord := 16#0100_0000;
      RED_ON_01 : DWord := 16#0800_0000;
      RED_ON_02 : DWord := 16#4000_0000;
      RED_ON_03 : DWord := 16#0002_0000;
      RED_ON_04 : DWord := 16#0010_0000;
      RED_ON_05 : DWord := 16#0080_0000;
      PART_00 : Int := 7;
      PART_01 : Int := 3;
      PART_02 : Int := 6;
      PART_03 : Int := 2;
      PART_04 : Int := 5;
      PART_05 : Int := 1;
   END_VAR
BEGIN
   IF #animator THEN
       "Stack_Light.Off"(part_number := #part_number,
                         stack_light := #stack_light);
       RETURN;
   END_IF;
   "Stack_Light.Red"(part_number := #part_number,
                     stack_light := #stack_light);
END_FUNCTION

FUNCTION "Stack_Light.Yellow" : Void   // FC329, SCL
{ S7_Optimized_Access := 'TRUE' }
VERSION : 0.1
   VAR_INPUT
      part_number : Int;
   END_VAR
   VAR_IN_OUT
      stack_light : DWord;
   END_VAR
   VAR CONSTANT
      YELLOW_ON_00 : DWord := 16#0200_0000;
      YELLOW_ON_01 : DWord := 16#1000_0000;
      YELLOW_ON_02 : DWord := 16#8000_0000;
      YELLOW_ON_03 : DWord := 16#0004_0000;
      YELLOW_ON_04 : DWord := 16#0020_0000;
      YELLOW_ON_05 : DWord := 16#0000_0100;
      PART_00 : Int := 7;
      PART_01 : Int := 3;
      PART_02 : Int := 6;
      PART_03 : Int := 2;
      PART_04 : Int := 5;
      PART_05 : Int := 1;
   END_VAR
BEGIN
   CASE #part_number OF
       #PART_00:
           #stack_light := #stack_light OR #YELLOW_ON_00;
       #PART_01:
           #stack_light := #stack_light OR #YELLOW_ON_01;
       #PART_02:
           #stack_light := #stack_light OR #YELLOW_ON_02;
       #PART_03:
           #stack_light := #stack_light OR #YELLOW_ON_03;
       #PART_04:
           #stack_light := #stack_light OR #YELLOW_ON_04;
       #PART_05:
           #stack_light := #stack_light OR #YELLOW_ON_05;
       ELSE
           ;
   END_CASE;
END_FUNCTION

FUNCTION "Stack_Light.Red" : Void   // FC330, SCL
{ S7_Optimized_Access := 'TRUE' }
VERSION : 0.1
   VAR_INPUT
      part_number : Int;
   END_VAR
   VAR_IN_OUT
      stack_light : DWord;
   END_VAR
   VAR CONSTANT
      RED_ON_00 : DWord := 16#0100_0000;
      RED_ON_01 : DWord := 16#0800_0000;
      RED_ON_02 : DWord := 16#4000_0000;
      RED_ON_03 : DWord := 16#0002_0000;
      RED_ON_04 : DWord := 16#0010_0000;
      RED_ON_05 : DWord := 16#0080_0000;
      PART_00 : Int := 7;
      PART_01 : Int := 3;
      PART_02 : Int := 6;
      PART_03 : Int := 2;
      PART_04 : Int := 5;
      PART_05 : Int := 1;
   END_VAR
BEGIN
   CASE #part_number OF
       #PART_00:
           #stack_light := #stack_light OR #RED_ON_00;
       #PART_01:
           #stack_light := #stack_light OR #RED_ON_01;
       #PART_02:
           #stack_light := #stack_light OR #RED_ON_02;
       #PART_03:
           #stack_light := #stack_light OR #RED_ON_03;
       #PART_04:
           #stack_light := #stack_light OR #RED_ON_04;
       #PART_05:
           #stack_light := #stack_light OR #RED_ON_05;
       ELSE
           ;
   END_CASE;
END_FUNCTION

FUNCTION "Stack_Light.Off" : Void   // FC331, SCL
{ S7_Optimized_Access := 'TRUE' }
VERSION : 0.1
   VAR_INPUT
      part_number : Int;
   END_VAR
   VAR_IN_OUT
      stack_light : DWord;
   END_VAR
   VAR CONSTANT
      GREEN_ON_00 : DWord := 16#0400_0000;
      RED_ON_00 : DWord := 16#0100_0000;
      YELLOW_ON_00 : DWord := 16#0200_0000;
      GREEN_ON_01 : DWord := 16#2000_0000;
      RED_ON_01 : DWord := 16#0800_0000;
      YELLOW_ON_01 : DWord := 16#1000_0000;
      GREEN_ON_02 : DWord := 16#0001_0000;
      RED_ON_02 : DWord := 16#4000_0000;
      YELLOW_ON_02 : DWord := 16#8000_0000;
      GREEN_ON_03 : DWord := 16#0008_0000;
      YELLOW_ON_03 : DWord := 16#0004_0000;
      RED_ON_03 : DWord := 16#0002_0000;
      GREEN_ON_04 : DWord := 16#0040_0000;
      RED_ON_04 : DWord := 16#0010_0000;
      YELLOW_ON_04 : DWord := 16#0020_0000;
      GREEN_ON_05 : DWord := 16#0000_0200;
      RED_ON_05 : DWord := 16#0080_0000;
      YELLOW_ON_05 : DWord := 16#0000_0100;
      PART_00 : Int := 7;
      PART_01 : Int := 3;
      PART_02 : Int := 6;
      PART_03 : Int := 2;
      PART_04 : Int := 5;
      PART_05 : Int := 1;
   END_VAR
BEGIN
   CASE #part_number OF
       #PART_00:
           #stack_light := #stack_light AND NOT #RED_ON_00;
           #stack_light := #stack_light AND NOT #YELLOW_ON_00;
           #stack_light := #stack_light AND NOT #GREEN_ON_00;
       #PART_01:
           #stack_light := #stack_light AND NOT #RED_ON_01;
           #stack_light := #stack_light AND NOT #YELLOW_ON_01;
           #stack_light := #stack_light AND NOT #GREEN_ON_01;
       #PART_02:
           #stack_light := #stack_light AND NOT #RED_ON_02;
           #stack_light := #stack_light AND NOT #YELLOW_ON_02;
           #stack_light := #stack_light AND NOT #GREEN_ON_02;
       #PART_03:
           #stack_light := #stack_light AND NOT #RED_ON_03;
           #stack_light := #stack_light AND NOT #YELLOW_ON_03;
           #stack_light := #stack_light AND NOT #GREEN_ON_03;
       #PART_04:
           #stack_light := #stack_light AND NOT #RED_ON_04;
           #stack_light := #stack_light AND NOT #YELLOW_ON_04;
           #stack_light := #stack_light AND NOT #GREEN_ON_04;
       #PART_05:
           #stack_light := #stack_light AND NOT #RED_ON_05;
           #stack_light := #stack_light AND NOT #YELLOW_ON_05;
           #stack_light := #stack_light AND NOT #GREEN_ON_05;
       ELSE
           ;
   END_CASE;
END_FUNCTION

// folder: Stations

FUNCTION_BLOCK "Button Parameters"   // FB12, SCL
{ S7_Optimized_Access := 'TRUE' }
VERSION : 0.1
   VAR_INPUT
      pnLib : "Recipe: PN Text Library";
   END_VAR
   VAR_IN_OUT
      stns : "Station: All Stations";
   END_VAR
   VAR
      placeHolder : Bool;
   END_VAR
   VAR_TEMP
      pBtn : Int;
      pStn : Int;
   END_VAR
BEGIN
   REGION "FOR EACH STATION"
       FOR #pStn := 0 TO "STATION_COUNT" DO

           REGION "ON CODE CHANGE"
               IF #stns.stn[#pStn].wipCmpts.flags.new_part_number THEN

                   REGION "FOR EACH BUTTON"
                       FOR #pBtn := 0 TO "BUTTON_COUNT" DO

                           REGION "LOAD PARAMETERS"
                               "Load Button Parameters OP"(pnGood := #stns.stn[#pStn].wipCmpts.flags.part_number_good[#pBtn],
                                                           btnConfig := #stns.stn[#pStn].kp8Config.btn[#pBtn]);
                           END_REGION

                       END_FOR;
                   END_REGION

               END_IF;
           END_REGION

       END_FOR;
   END_REGION
END_FUNCTION_BLOCK

FUNCTION "Load Button Parameters OP" : Void   // FC2, SCL
{ S7_Optimized_Access := 'TRUE' }
VERSION : 0.1
   VAR_INPUT
      pnGood : Bool;
   END_VAR
   VAR_IN_OUT
      btnConfig : "KP8 Driver: Parameters: 1 Button";
   END_VAR
BEGIN
   REGION "ON GOOD PN"
       IF #pnGood THEN

           REGION "ACTIVATE BUTTON"
               #btnConfig.activate := TRUE;
               #btnConfig.cOff := 'green';
               #btnConfig.cOn1 := 'yellow';
               #btnConfig.cOn2 := '';
               #btnConfig.flash := FALSE;
               #btnConfig.group := 0;
               #btnConfig.mode := TRUE;
           END_REGION

       END_IF;
   END_REGION

   REGION "ON BAD PN"
       IF NOT #pnGood THEN

